               Strg_TO_Chars(Strg:= CONCAT_STRING(IN1 := #TMP_strTemp ,IN2 := DINT_TO_STRING(#IN_rgtStatusMarkers[#TMP_dMarkerIndex].dStatus)),
                         pChars:=#TMP_dIndex,
                         Cnt=>#TMP_uiNumChar,
                         Chars:=#AUX_rgcStatusTelegram);
               #TMP_dIndex+=#TMP_uiNumChar;

               #AUX_rgcStatusTelegram[#TMP_dIndex] := #STRSEPARATOR;
               #TMP_dIndex+=1;
           END_IF;

           IF (#IN_rgtStatusMarkers[#TMP_dMarkerIndex].dMarkerActualStatus <> #AUX_rgtStatusMarkers[#TMP_dMarkerIndex].dMarkerActualStatus) OR (#AUX_xResendAllStatus) THEN

               #AUX_rgtStatusMarkers[#TMP_dMarkerIndex].dMarkerActualStatus := #IN_rgtStatusMarkers[#TMP_dMarkerIndex].dMarkerActualStatus;        

               #TMP_strTemp := CONCAT_STRING(IN1 := #STRSTATUSMARKACTSTATUS ,IN2 := #TMP_strMarkerIndex);
               #TMP_strTemp := CONCAT_STRING(IN1 := #TMP_strTemp ,IN2 := '=');

               Strg_TO_Chars(Strg:= CONCAT_STRING(IN1 := #TMP_strTemp ,IN2 := DINT_TO_STRING(#IN_rgtStatusMarkers[#TMP_dMarkerIndex].dMarkerActualStatus)),
                         pChars:=#TMP_dIndex,
                         Cnt=>#TMP_uiNumChar,
                         Chars:=#AUX_rgcStatusTelegram);
               #TMP_dIndex+=#TMP_uiNumChar;

               #AUX_rgcStatusTelegram[#TMP_dIndex] := #STRSEPARATOR;
               #TMP_dIndex+=1;
           END_IF;*)


       END_FOR;

       END_REGION BPS_STATUS_TELEGRAM_MARKERS

       REGION BPS_STATUS_TELEGRAM_YCUTS

       FOR #TMP_dYCutIndex := 0 TO "DMAXYCUTBRIDGE_IND" DO

           #TMP_strYCutIndex := DINT_TO_STRING(#TMP_dYCutIndex + 1);   

           #TMP_strYCutIndex := DELETE(IN:=#TMP_strYCutIndex, L:=1, P:=1);

           //Prepare position information
           #TMP_strYCut := CONCAT_STRING(IN1 := #STRSTATUSYCUT ,IN2 := #TMP_strYCutIndex);

           IF (#IN_rgtStatusYCuts[#TMP_dYCutIndex].dBridgeStatus <> #AUX_rgtStatusYCuts[#TMP_dYCutIndex].dBridgeStatus) OR (#AUX_xResendAllStatus) THEN

               #AUX_rgtStatusYCuts[#TMP_dYCutIndex].dBridgeStatus := #IN_rgtStatusYCuts[#TMP_dYCutIndex].dBridgeStatus;        

               #TMP_strTemp := CONCAT_STRING(IN1 := #TMP_strYCut ,IN2 := #STRSTATUSYCUTSTATUS);

               Strg_TO_Chars(Strg:= CONCAT_STRING(IN1 := #TMP_strTemp ,IN2 := DINT_TO_STRING(#IN_rgtStatusYCuts[#TMP_dYCutIndex].dBridgeStatus)),
                         pChars:=#TMP_dIndex,
                         Cnt=>#TMP_uiNumChar,
                         Chars:=#AUX_rgcStatusTelegram);
               #TMP_dIndex+=#TMP_uiNumChar;

               #AUX_rgcStatusTelegram[#TMP_dIndex] := #STRSEPARATOR;
               #TMP_dIndex+=1;
           END_IF;

           IF (#IN_rgtStatusYCuts[#TMP_dYCutIndex].dDistanceSnapRoll_cmm <> #AUX_rgtStatusYCuts[#TMP_dYCutIndex].dDistanceSnapRoll_cmm) OR (#AUX_xResendAllStatus) THEN

               #AUX_rgtStatusYCuts[#TMP_dYCutIndex].dDistanceSnapRoll_cmm := #IN_rgtStatusYCuts[#TMP_dYCutIndex].dDistanceSnapRoll_cmm;        

               #TMP_strTemp := CONCAT_STRING(IN1 := #TMP_strYCut ,IN2 := #STRSTATUSYCUTSDISTSNAP);

               Strg_TO_Chars(Strg:= CONCAT_STRING(IN1 := #TMP_strTemp ,IN2 := DINT_TO_STRING(#IN_rgtStatusYCuts[#TMP_dYCutIndex].dDistanceSnapRoll_cmm)),
                         pChars:=#TMP_dIndex,
                         Cnt=>#TMP_uiNumChar,
                         Chars:=#AUX_rgcStatusTelegram);
               #TMP_dIndex+=#TMP_uiNumChar;

               #AUX_rgcStatusTelegram[#TMP_dIndex] := #STRSEPARATOR;
               #TMP_dIndex+=1;
           END_IF;


           FOR #TMP_dYCutHeadIndex := 0 TO "DMAXYHEADS_IND" DO

               #TMP_strHeadIndex := DINT_TO_STRING(#TMP_dYCutHeadIndex + 1);
               #TMP_strHeadIndex := DELETE(IN:=#TMP_strHeadIndex, L:= 1, P:=1);

               IF (#IN_rgtStatusYCuts[#TMP_dYCutIndex].rgdPosition_cmm[#TMP_dYCutHeadIndex] <> #AUX_rgtStatusYCuts[#TMP_dYCutIndex].rgdPosition_cmm[#TMP_dYCutHeadIndex]) OR (#AUX_xResendAllStatus) THEN

                   #AUX_rgtStatusYCuts[#TMP_dYCutIndex].rgdPosition_cmm[#TMP_dYCutHeadIndex] := #IN_rgtStatusYCuts[#TMP_dYCutIndex].rgdPosition_cmm[#TMP_dYCutHeadIndex];

                   #TMP_strTemp := CONCAT_STRING(IN1 := #TMP_strYCut ,IN2 := #STRSTATUSYCUTPOS);
                   #TMP_strTemp := CONCAT_STRING(IN1 := #TMP_strTemp, IN2 := #TMP_strHeadIndex);
                   #TMP_strTemp := CONCAT_STRING(IN1 := #TMP_strTemp,IN2 := '=');

                   Strg_TO_Chars(Strg:= CONCAT_STRING(IN1 := #TMP_strTemp ,IN2 := DINT_TO_STRING(#IN_rgtStatusYCuts[#TMP_dYCutIndex].rgdPosition_cmm[#TMP_dYCutHeadIndex])),
                         pChars:=#TMP_dIndex,
                         Cnt=>#TMP_uiNumChar,
                         Chars:=#AUX_rgcStatusTelegram);
                   #TMP_dIndex+=#TMP_uiNumChar;

                   #AUX_rgcStatusTelegram[#TMP_dIndex] := #STRSEPARATOR;
                   #TMP_dIndex+=1;
               END_IF;

               IF (#IN_rgtStatusYCuts[#TMP_dYCutIndex].rgxFireON[#TMP_dYCutHeadIndex] <> #AUX_rgtStatusYCuts[#TMP_dYCutIndex].rgxFireON[#TMP_dYCutHeadIndex]) OR (#AUX_xResendAllStatus) THEN

                   #AUX_rgtStatusYCuts[#TMP_dYCutIndex].rgxFireON[#TMP_dYCutHeadIndex] := #IN_rgtStatusYCuts[#TMP_dYCutIndex].rgxFireON[#TMP_dYCutHeadIndex];

                   #TMP_strTemp := CONCAT_STRING(IN1 := #TMP_strYCut ,IN2 := #STRSTATUSYCUTFIRE);
                   #TMP_strTemp := CONCAT_STRING(IN1 := #TMP_strTemp, IN2 := #TMP_strHeadIndex);
                   #TMP_strTemp := CONCAT_STRING(IN1 := #TMP_strTemp,IN2 := '=');

                   Strg_TO_Chars(Strg:= CONCAT_STRING(IN1 := #TMP_strTemp ,IN2 := DINT_TO_STRING(BOOL_TO_DINT(#IN_rgtStatusYCuts[#TMP_dYCutIndex].rgxFireON[#TMP_dYCutHeadIndex]))),
                         pChars:=#TMP_dIndex,
                         Cnt=>#TMP_uiNumChar,
                         Chars:=#AUX_rgcStatusTelegram);
                   #TMP_dIndex+=#TMP_uiNumChar;

                   #AUX_rgcStatusTelegram[#TMP_dIndex] := #STRSEPARATOR;
                   #TMP_dIndex+=1;
               END_IF;

               IF (#IN_rgtStatusYCuts[#TMP_dYCutIndex].rgxArmON[#TMP_dYCutHeadIndex] <> #AUX_rgtStatusYCuts[#TMP_dYCutIndex].rgxArmON[#TMP_dYCutHeadIndex]) OR (#AUX_xResendAllStatus) THEN

                   #AUX_rgtStatusYCuts[#TMP_dYCutIndex].rgxArmON[#TMP_dYCutHeadIndex] := #IN_rgtStatusYCuts[#TMP_dYCutIndex].rgxArmON[#TMP_dYCutHeadIndex];

                   #TMP_strTemp := CONCAT_STRING(IN1 := #TMP_strYCut ,IN2 := #STRSTATUSYCUTARM);
                   #TMP_strTemp := CONCAT_STRING(IN1 := #TMP_strTemp, IN2 := #TMP_strHeadIndex);
                   #TMP_strTemp := CONCAT_STRING(IN1 := #TMP_strTemp,IN2 := '=');

                   Strg_TO_Chars(Strg:= CONCAT_STRING(IN1 := #TMP_strTemp ,IN2 := DINT_TO_STRING(BOOL_TO_DINT(#IN_rgtStatusYCuts[#TMP_dYCutIndex].rgxArmON[#TMP_dYCutHeadIndex]))),
                         pChars:=#TMP_dIndex,
                         Cnt=>#TMP_uiNumChar,
                         Chars:=#AUX_rgcStatusTelegram);
                   #TMP_dIndex+=#TMP_uiNumChar;

                   #AUX_rgcStatusTelegram[#TMP_dIndex] := #STRSEPARATOR;
                   #TMP_dIndex+=1;
               END_IF;

               IF (#IN_rgtStatusYCuts[#TMP_dYCutIndex].rgxHeadProdOn[#TMP_dYCutHeadIndex] <> #AUX_rgtStatusYCuts[#TMP_dYCutIndex].rgxHeadProdOn[#TMP_dYCutHeadIndex]) OR (#AUX_xResendAllStatus) THEN

                   #AUX_rgtStatusYCuts[#TMP_dYCutIndex].rgxHeadProdOn[#TMP_dYCutHeadIndex] := #IN_rgtStatusYCuts[#TMP_dYCutIndex].rgxHeadProdOn[#TMP_dYCutHeadIndex];

                   #TMP_strTemp := CONCAT_STRING(IN1 := #TMP_strYCut ,IN2 := #STRSTATUSYCUTPROD);
                   #TMP_strTemp := CONCAT_STRING(IN1 := #TMP_strTemp, IN2 := #TMP_strHeadIndex);
                   #TMP_strTemp := CONCAT_STRING(IN1 := #TMP_strTemp,IN2 := '=');

                   Strg_TO_Chars(Strg:= CONCAT_STRING(IN1 := #TMP_strTemp ,IN2 := DINT_TO_STRING(BOOL_TO_DINT(#IN_rgtStatusYCuts[#TMP_dYCutIndex].rgxHeadProdOn[#TMP_dYCutHeadIndex]))),
                         pChars:=#TMP_dIndex,
                         Cnt=>#TMP_uiNumChar,
                         Chars:=#AUX_rgcStatusTelegram);
                   #TMP_dIndex+=#TMP_uiNumChar;

                   #AUX_rgcStatusTelegram[#TMP_dIndex] := #STRSEPARATOR;
                   #TMP_dIndex+=1;
               END_IF;

           END_FOR;


       END_FOR;

      // #AUX_xResendAllStatus := FALSE;


       END_REGION BPS_STATUS_TELEGRAM_YCUTS


       #AUX_rgcStatusTelegram[#TMP_dIndex] := #STR_CR;
       #TMP_dIndex+=1;

       #AUX_rgcStatusTelegram[#TMP_dIndex] := #STR_LF;

       #AUX_dStatusTelegramNumByte := #TMP_dIndex + 1;

       IF #AUX_dStatusTelegramCounter >= #DMAXTELEGRAMCOUNTER THEN
           #AUX_dStatusTelegramCounter := 1;
       ELSE
           #AUX_dStatusTelegramCounter += 1;
       END_IF;

       IF (((#IN_xBPSServerA) AND (#IN_tStatusGeneral.dExtOptSelected = 1)) OR
           ((NOT #IN_xBPSServerA) AND (#IN_tStatusGeneral.dExtOptSelected = 2))) THEN

           IF #AUX_dStatusServerCounter >= #DMAXTELEGRAMCOUNTER THEN
               #AUX_dStatusServerCounter := 1;
           ELSE
               #AUX_dStatusServerCounter += 1;
           END_IF;

       END_IF;    
       #ST_xStatusTelegramAvail := TRUE;

   END_IF;





   END_REGION BPS_STATUS_TELEGRAM

   REGION BPS_SEND_INFORMATION

   //Initialize connection data in case of reset
   IF #IN_xGeneralReset THEN

       #AUX_tConnData.InterfaceId := #IN_tInterfaceID;
       #AUX_tConnData.ID := #IN_tID;
       #AUX_tConnData.ConnectionType := #BCONNTYPE;
       #AUX_tConnData.ActiveEstablished := TRUE;
       #AUX_tConnData.RemoteAddress := #IN_tRemoteAddress;
       #AUX_tConnData.RemotePort := #IN_uiRemotePort;
       #AUX_tConnData.LocalPort := 0;

       //Reset della fasi
       #TMP_dwValue := 0;
       SCATTER(IN:=#TMP_dwValue,
               OUT=>#tPhasesNetwork);

       //Reset others data
       #ST_xRetrySendTelegram := FALSE;
       #AUX_dSendTelegramNumByte := 0;
       #TMP_cValue := ' ';

       FILL_BLK(IN:=#TMP_cValue,
                COUNT:=DINT_TO_ULINT(#DSENDTELEGRAMSIZE),
                OUT=>#AUX_rgcSendTelegram[0]);


   END_IF;

   #AUX_xResetSendConnection := #IN_xGeneralReset OR (#FB_TSend.s_TDIAG_Status.State <> b#16#04 AND #IN_xResetAlarms);


   IF NOT #ST_xPhasesInProgress AND #IN_xThisPLCActive AND
           (#ST_xPlateTelegramAvail OR 
           #ST_xStatusTelegramAvail OR 
           #ST_xDefectTelegramAvail OR 
           #ST_xRibbonTelegramAvail OR 
           #ST_xEventsTelegramAvail OR
           #ST_xRibbonTelegramAvail OR 
           #ST_xRetrySendTelegram) THEN

       IF NOT #ST_xRetrySendTelegram THEN

           //Fill the send buffer with the status telegram and plate
           #AUX_dSendTelegramNumByte := 0;

           IF #ST_xPlateTelegramAvail THEN

               MOVE_BLK(IN:=#AUX_rgcPlateTelegram[0],
                        COUNT:=DINT_TO_ULINT(#AUX_dPlateTelegramNumByte),
                        OUT=>#AUX_rgcSendTelegram[0]);

               #AUX_dSendTelegramNumByte:= #AUX_dPlateTelegramNumByte;

               #ST_xPlateTelegramAvail := FALSE;
               #AUX_xResendAllPlate := FALSE;
           ELSIF #ST_xStatusTelegramAvail THEN

               MOVE_BLK(IN := #AUX_rgcStatusTelegram[0],
                        COUNT := DINT_TO_ULINT(#AUX_dStatusTelegramNumByte),
                        OUT => #AUX_rgcSendTelegram[0]);

               #AUX_dSendTelegramNumByte := #AUX_dStatusTelegramNumByte;

               #ST_xStatusTelegramAvail := FALSE;
               #AUX_xResendAllStatus := FALSE;


           ELSIF #ST_xDefectTelegramAvail THEN

               MOVE_BLK(IN:=#AUX_rgcDefectTelegram[0],
                        COUNT:=DINT_TO_ULINT(#AUX_dDefectTelegramNumByte),
                        OUT=>#AUX_rgcSendTelegram[0]);

               #AUX_dSendTelegramNumByte:= #AUX_dDefectTelegramNumByte;

               #ST_xDefectTelegramAvail := FALSE;

           ELSIF #ST_xEventsTelegramAvail THEN

               MOVE_BLK(IN:=#AUX_rgcEventsTelegram[0],
                        COUNT:=DINT_TO_ULINT(#AUX_dEventsTelegramNumByte),
                        OUT=>#AUX_rgcSendTelegram[0]);

               #AUX_dSendTelegramNumByte:= #AUX_dEventsTelegramNumByte;

               #ST_xEventsTelegramAvail := FALSE;

           ELSIF #ST_xRibbonTelegramAvail THEN

               MOVE_BLK(IN:=#AUX_rgcRibbonTelegram[0],
                        COUNT:=DINT_TO_ULINT(#AUX_dRibbonTelegramNumByte),
                        OUT=>#AUX_rgcSendTelegram[0]);

               #AUX_dSendTelegramNumByte:= #AUX_dRibbonTelegramNumByte;

               #ST_xRibbonTelegramAvail := FALSE;

          ELSIF #ST_xStatusTelegramAvail THEN

               MOVE_BLK(IN:=#AUX_rgcStatusTelegram[0],
                        COUNT:=DINT_TO_ULINT(#AUX_dStatusTelegramNumByte),
                        OUT=>#AUX_rgcSendTelegram[0]);

               #AUX_dSendTelegramNumByte:= #AUX_dStatusTelegramNumByte;

               #ST_xStatusTelegramAvail := FALSE;
               #AUX_xResendAllStatus := FALSE;
           END_IF;

       END_IF;


       #tPhasesNetwork.xSendBufferInProgress := TRUE; 

   END_IF;


   #FB_TSend(REQ:=#tPhasesNetwork.xSendBufferInProgress,
             CONT:=#IN_xThisPLCActive,
             LEN:=DINT_TO_UDINT(#AUX_dSendTelegramNumByte),
             CONNECT:=#AUX_tConnData,
             DATA:=#AUX_rgcSendTelegram,
             COM_RST:=#AUX_xResetSendConnection);


   //Manage send feedback
   IF #tPhasesNetwork.xSendBufferInProgress AND 
                                           (#FB_TSend.DONE OR
                                           #FB_TSend.ERROR OR 
                                           NOT #FB_TSend.BUSY) THEN

       #tPhasesNetwork.xSendBufferInProgress := FALSE;
       #tPhasesNetwork.xEndSendBufferInProgress := TRUE;
       #ST_xRetrySendTelegram := FALSE;
       IF NOT #FB_TSend.DONE THEN

           #ST_xRetrySendTelegram := TRUE;

       END_IF;

   ELSE

       #tPhasesNetwork.xEndSendBufferInProgress := FALSE;
   END_IF;

   //Calculate phase in progress
   GATHER(IN:=#tPhasesNetwork,
          OUT=>#TMP_dwValue);

   IF #TMP_dwValue <> 0 THEN
       #ST_xPhasesInProgress := TRUE;
   ELSE
       #ST_xPhasesInProgress := FALSE;
   END_IF;




   END_REGION BPS_SEND_INFORMATION

   REGION BPS_RECEIVE_INFORMATION

   #FB_TRecv(EN_R:=#IN_xThisPLCActive,
             CONT:=#IN_xThisPLCActive,
             LEN:=0,
             ADHOC:=TRUE,
             CONNECT:=#AUX_tConnData,
             DATA:=#AUX_rgcRecvTelegram,
             COM_RST:=#AUX_xResetSendConnection);

   IF #FB_TRecv.DONE THEN

       IF (#FB_TRecv.RCVD_LEN > 0) AND (UDINT_TO_DINT(#FB_TRecv.RCVD_LEN) + #AUX_dNumByteRecvBuffer < #DRECVBUFFERSIZE) THEN

           //Copy the received data
           #TMP_iRetVal := MOVE_BLK_VARIANT(SRC:=#AUX_rgcRecvTelegram, COUNT:=#FB_TRecv.RCVD_LEN, SRC_INDEX:=0, DEST_INDEX:=#AUX_dNumByteRecvBuffer, DEST=>#AUX_rgcRecvBuffer);
           #AUX_dNumByteRecvBuffer += UDINT_TO_DINT(#FB_TRecv.RCVD_LEN);

       END_IF;

   END_IF;

   //Analyze telegrams 
   FOR #TMP_dIndex := 0 TO #AUX_dNumByteRecvBuffer - 2 DO

       IF (#AUX_rgcRecvBuffer[#TMP_dIndex] = #STR_CR) AND (#AUX_rgcRecvBuffer[#TMP_dIndex + 1] = #STR_LF) THEN

           //End of packet found. Move the data to a string
           #TMP_iRetVal := MOVE_BLK_VARIANT(SRC:=#AUX_rgcRecvBuffer, COUNT:= DINT_TO_UDINT(#TMP_dIndex) + 2 , SRC_INDEX:= 0, DEST_INDEX:= 0, DEST=>#AUX_rgcAnalyzedTelegram);

           IF (#TMP_dIndex + 2) < #AUX_dNumByteRecvBuffer THEN
               #TMP_iRetVal := MOVE_BLK_VARIANT(SRC:=#AUX_rgcRecvBuffer, COUNT:=DINT_TO_UDINT(#AUX_dNumByteRecvBuffer - (#TMP_dIndex + 2))   , SRC_INDEX:= #TMP_dIndex + 2 , DEST_INDEX:= 0, DEST=>#AUX_rgcRecvBuffer);
           ELSE
               #AUX_dNumByteRecvBuffer := 0;
           END_IF;
           #TMP_udCountString := 0;
           #TMP_udPosition := 0;
           #TMP_cSeparator := #STRSEPARATOR;

           #TMP_cEndSeparator := #STR_LF;
           //Split the telegram and manage it
           #TMP_iRetVal := SPLIT(Mode:=0, RecSeparator:=#TMP_cSeparator, EndSeparator:=#TMP_cEndSeparator, SrcArray:=#AUX_rgcAnalyzedTelegram, Count=>#TMP_udCountString, DstStruct:=#AUX_rgstrMessageString, Position:=#TMP_udPosition);

   REGION BPS_RECEIVE_EVENT 
           //Check the received message 'D'
           IF (#AUX_rgstrMessageString[0] = CHAR_TO_STRING(#STREVENTSTELEGRAMID)) AND (#TMP_udCountString = 16) THEN

               //Event code
               #TMP_cSeparator := '=';
               #TMP_uiCount := 0;


               Strg_TO_Chars(Strg:=#AUX_rgstrMessageString[2],
                             pChars:=0,
                             Cnt=>#TMP_uiCount,
                             Chars:=#AUX_rgcMetaData);
               #AUX_rgcMetaData[#TMP_uiCount] := #STR_LF;
               #TMP_udPosition := 0;
               #TMP_iRetVal := SPLIT(  Mode:=0, 
                                       RecSeparator:=#TMP_cSeparator, 
                                       EndSeparator:=#TMP_cEndSeparator, 
                                       SrcArray:=#AUX_rgcMetaData, 
                                       Count=>#TMP_udCountString, 
                                       DstStruct:=#AUX_rgstrSingleMexString, 
                                       Position:=#TMP_udPosition);
               IF ( #TMP_udCountString = 2) AND #AUX_rgstrSingleMexString[0] = 'Cd' THEN
                   #AUX_tRecvMessage.dCodeEvent := STRING_TO_DINT(#AUX_rgstrSingleMexString[1]);
               ELSE 
                   #AUX_tRecvMessage.dCodeEvent := 0;
               END_IF;

               //Ident
               #TMP_cSeparator := '=';
               #TMP_uiCount := 0;
               Strg_TO_Chars(Strg:=#AUX_rgstrMessageString[4],
                             pChars:=0,
                             Cnt=>#TMP_uiCount,
                             Chars:=#AUX_rgcMetaData);
               #AUX_rgcMetaData[#TMP_uiCount] := #STR_LF;
               #TMP_udPosition := 0;
               #TMP_iRetVal := SPLIT(  Mode:=0, 
                                       RecSeparator:=#TMP_cSeparator, 
                                       EndSeparator:=#TMP_cEndSeparator, 
                                       SrcArray:=#AUX_rgcMetaData, 
                                       Count=>#TMP_udCountString, 
                                       DstStruct:=#AUX_rgstrSingleMexString, 
                                       Position:=#TMP_udPosition);
               IF ( #TMP_udCountString = 2) AND #AUX_rgstrSingleMexString[0] = 'Id' THEN
                   #AUX_tRecvMessage.strIdent := #AUX_rgstrSingleMexString[1];
               ELSE 
                   #AUX_tRecvMessage.strIdent := '';
               END_IF;

               //Data 1
               #TMP_cSeparator := '=';
               #TMP_uiCount := 0;
               Strg_TO_Chars(Strg:=#AUX_rgstrMessageString[5],
                             pChars:=0,
                             Cnt=>#TMP_uiCount,
                             Chars:=#AUX_rgcMetaData);
               #AUX_rgcMetaData[#TMP_uiCount] := #STR_LF;
               #TMP_udPosition := 0;
               #TMP_iRetVal := SPLIT(  Mode:=0, 
                                       RecSeparator:=#TMP_cSeparator, 
                                       EndSeparator:=#TMP_cEndSeparator, 
                                       SrcArray:=#AUX_rgcMetaData, 
                                       Count=>#TMP_udCountString, 
                                       DstStruct:=#AUX_rgstrSingleMexString, 
                                       Position:=#TMP_udPosition);
               IF ( #TMP_udCountString = 2) AND #AUX_rgstrSingleMexString[0] = 'D1' THEN
                   #AUX_tRecvMessage.dEvent1 := STRING_TO_DINT(#AUX_rgstrSingleMexString[1]);
               ELSE 
                   #AUX_tRecvMessage.dEvent1 := 0;
               END_IF;

               //Data 2
               #TMP_cSeparator := '=';
               #TMP_uiCount := 0;
               Strg_TO_Chars(Strg:=#AUX_rgstrMessageString[6],
                             pChars:=0,
                             Cnt=>#TMP_uiCount,
                             Chars:=#AUX_rgcMetaData);
               #AUX_rgcMetaData[#TMP_uiCount] := #STR_LF;
               #TMP_udPosition := 0;
               #TMP_iRetVal := SPLIT(  Mode:=0, 
                                       RecSeparator:=#TMP_cSeparator, 
                                       EndSeparator:=#TMP_cEndSeparator, 
                                       SrcArray:=#AUX_rgcMetaData, 
                                       Count=>#TMP_udCountString, 
                                       DstStruct:=#AUX_rgstrSingleMexString, 
                                       Position:=#TMP_udPosition);
               IF ( #TMP_udCountString = 2) AND #AUX_rgstrSingleMexString[0] = 'D2' THEN
                   #AUX_tRecvMessage.dEvent2 := STRING_TO_DINT(#AUX_rgstrSingleMexString[1]);
               ELSE 
                   #AUX_tRecvMessage.dEvent2 := 0;
               END_IF;

               //Data 3
               #TMP_cSeparator := '=';
               #TMP_uiCount := 0;
               Strg_TO_Chars(Strg:=#AUX_rgstrMessageString[7],
                             pChars:=0,
                             Cnt=>#TMP_uiCount,
                             Chars:=#AUX_rgcMetaData);
               #AUX_rgcMetaData[#TMP_uiCount] := #STR_LF;
               #TMP_udPosition := 0;
               #TMP_iRetVal := SPLIT(  Mode:=0, 
                                       RecSeparator:=#TMP_cSeparator, 
                                       EndSeparator:=#TMP_cEndSeparator, 
                                       SrcArray:=#AUX_rgcMetaData, 
                                       Count=>#TMP_udCountString, 
                                       DstStruct:=#AUX_rgstrSingleMexString, 
                                       Position:=#TMP_udPosition);
               IF ( #TMP_udCountString = 2) AND #AUX_rgstrSingleMexString[0] = 'D3' THEN
                   #AUX_tRecvMessage.dEvent3 := STRING_TO_DINT(#AUX_rgstrSingleMexString[1]);
               ELSE 
                   #AUX_tRecvMessage.dEvent3 := 0;
               END_IF;

               //Data 4
               #TMP_cSeparator := '=';
               #TMP_uiCount := 0;
               Strg_TO_Chars(Strg:=#AUX_rgstrMessageString[8],
                             pChars:=0,
                             Cnt=>#TMP_uiCount,
                             Chars:=#AUX_rgcMetaData);
               #AUX_rgcMetaData[#TMP_uiCount] := #STR_LF;
               #TMP_udPosition := 0;
               #TMP_iRetVal := SPLIT(  Mode:=0, 
                                       RecSeparator:=#TMP_cSeparator, 
                                       EndSeparator:=#TMP_cEndSeparator, 
                                       SrcArray:=#AUX_rgcMetaData, 
                                       Count=>#TMP_udCountString, 
                                       DstStruct:=#AUX_rgstrSingleMexString, 
                                       Position:=#TMP_udPosition);
               IF ( #TMP_udCountString = 2) AND #AUX_rgstrSingleMexString[0] = 'D4' THEN
                   #AUX_tRecvMessage.dEvent4 := STRING_TO_DINT(#AUX_rgstrSingleMexString[1]);
               ELSE 
                   #AUX_tRecvMessage.dEvent4 := 0;
               END_IF;

               //Data 5
               #TMP_cSeparator := '=';
               #TMP_uiCount := 0;
               Strg_TO_Chars(Strg:=#AUX_rgstrMessageString[9],
                             pChars:=0,
                             Cnt=>#TMP_uiCount,
                             Chars:=#AUX_rgcMetaData);
               #AUX_rgcMetaData[#TMP_uiCount] := #STR_LF;
               #TMP_udPosition := 0;
               #TMP_iRetVal := SPLIT(  Mode:=0, 
                                       RecSeparator:=#TMP_cSeparator, 
                                       EndSeparator:=#TMP_cEndSeparator, 
                                       SrcArray:=#AUX_rgcMetaData, 
                                       Count=>#TMP_udCountString, 
                                       DstStruct:=#AUX_rgstrSingleMexString, 
                                       Position:=#TMP_udPosition);
               IF ( #TMP_udCountString = 2) AND #AUX_rgstrSingleMexString[0] = 'D5' THEN
                   #AUX_tRecvMessage.dEvent5 := STRING_TO_DINT(#AUX_rgstrSingleMexString[1]);
               ELSE 
                   #AUX_tRecvMessage.dEvent5 := 0;
               END_IF;

               //Data 6
               #TMP_cSeparator := '=';
               #TMP_uiCount := 0;
               Strg_TO_Chars(Strg:=#AUX_rgstrMessageString[10],
                             pChars:=0,
                             Cnt=>#TMP_uiCount,
                             Chars:=#AUX_rgcMetaData);
               #AUX_rgcMetaData[#TMP_uiCount] := #STR_LF;
               #TMP_udPosition := 0;
               #TMP_iRetVal := SPLIT(  Mode:=0, 
                                       RecSeparator:=#TMP_cSeparator, 
                                       EndSeparator:=#TMP_cEndSeparator, 
                                       SrcArray:=#AUX_rgcMetaData, 
                                       Count=>#TMP_udCountString, 
                                       DstStruct:=#AUX_rgstrSingleMexString, 
                                       Position:=#TMP_udPosition);
               IF ( #TMP_udCountString = 2) AND #AUX_rgstrSingleMexString[0] = 'D6' THEN
                   #AUX_tRecvMessage.dEvent6 := STRING_TO_DINT(#AUX_rgstrSingleMexString[1]);
               ELSE 
                   #AUX_tRecvMessage.dEvent6 := 0;
               END_IF;

               //Data 7
               #TMP_cSeparator := '=';
               #TMP_uiCount := 0;
               Strg_TO_Chars(Strg:=#AUX_rgstrMessageString[11],
                             pChars:=0,
                             Cnt=>#TMP_uiCount,
                             Chars:=#AUX_rgcMetaData);
               #AUX_rgcMetaData[#TMP_uiCount] := #STR_LF;
               #TMP_udPosition := 0;
               #TMP_iRetVal := SPLIT(  Mode:=0, 
                                       RecSeparator:=#TMP_cSeparator, 
                                       EndSeparator:=#TMP_cEndSeparator, 
                                       SrcArray:=#AUX_rgcMetaData, 
                                       Count=>#TMP_udCountString, 
                                       DstStruct:=#AUX_rgstrSingleMexString, 
                                       Position:=#TMP_udPosition);
               IF ( #TMP_udCountString = 2) AND #AUX_rgstrSingleMexString[0] = 'D7' THEN
                   #AUX_tRecvMessage.dEvent7 := STRING_TO_DINT(#AUX_rgstrSingleMexString[1]);
               ELSE 
                   #AUX_tRecvMessage.dEvent7 := 0;
               END_IF;

               //Data 8
               #TMP_cSeparator := '=';
               #TMP_uiCount := 0;
               Strg_TO_Chars(Strg:=#AUX_rgstrMessageString[12],
                             pChars:=0,
                             Cnt=>#TMP_uiCount,
                             Chars:=#AUX_rgcMetaData);
               #AUX_rgcMetaData[#TMP_uiCount] := #STR_LF;
               #TMP_udPosition := 0;
               #TMP_iRetVal := SPLIT(  Mode:=0, 
                                       RecSeparator:=#TMP_cSeparator, 
                                       EndSeparator:=#TMP_cEndSeparator, 
                                       SrcArray:=#AUX_rgcMetaData, 
                                       Count=>#TMP_udCountString, 
                                       DstStruct:=#AUX_rgstrSingleMexString, 
                                       Position:=#TMP_udPosition);
               IF ( #TMP_udCountString = 2) AND #AUX_rgstrSingleMexString[0] = 'D8' THEN
                   #AUX_tRecvMessage.dEvent8 := STRING_TO_DINT(#AUX_rgstrSingleMexString[1]);
               ELSE 
                   #AUX_tRecvMessage.dEvent8 := 0;
               END_IF;

               //Data 9
               #TMP_cSeparator := '=';
               #TMP_uiCount := 0;
               Strg_TO_Chars(Strg:=#AUX_rgstrMessageString[13],
                             pChars:=0,
                             Cnt=>#TMP_uiCount,
                             Chars:=#AUX_rgcMetaData);
               #AUX_rgcMetaData[#TMP_uiCount] := #STR_LF;
               #TMP_udPosition := 0;
               #TMP_iRetVal := SPLIT(  Mode:=0, 
                                       RecSeparator:=#TMP_cSeparator, 
                                       EndSeparator:=#TMP_cEndSeparator, 
                                       SrcArray:=#AUX_rgcMetaData, 
                                       Count=>#TMP_udCountString, 
                                       DstStruct:=#AUX_rgstrSingleMexString, 
                                       Position:=#TMP_udPosition);
               IF ( #TMP_udCountString = 2) AND #AUX_rgstrSingleMexString[0] = 'D9' THEN
                   #AUX_tRecvMessage.dEvent9 := STRING_TO_DINT(#AUX_rgstrSingleMexString[1]);
               ELSE 
                   #AUX_tRecvMessage.dEvent9 := 0;
               END_IF;

               //Data 10
               #TMP_cSeparator := '=';
               #TMP_uiCount := 0;
               Strg_TO_Chars(Strg:=#AUX_rgstrMessageString[14],
                             pChars:=0,
                             Cnt=>#TMP_uiCount,
                             Chars:=#AUX_rgcMetaData);
               #AUX_rgcMetaData[#TMP_uiCount] := #STR_LF;
               #TMP_udPosition := 0;
               #TMP_iRetVal := SPLIT(  Mode:=0, 
                                       RecSeparator:=#TMP_cSeparator, 
                                       EndSeparator:=#TMP_cEndSeparator, 
                                       SrcArray:=#AUX_rgcMetaData, 
                                       Count=>#TMP_udCountString, 
                                       DstStruct:=#AUX_rgstrSingleMexString, 
                                       Position:=#TMP_udPosition);
               IF ( #TMP_udCountString = 2) AND #AUX_rgstrSingleMexString[0] = 'D10' THEN
                   #AUX_tRecvMessage.dEvent10 := STRING_TO_DINT(#AUX_rgstrSingleMexString[1]);
               ELSE 
                   #AUX_tRecvMessage.dEvent10 := 0;
               END_IF;

               "RP_AddMessageV2"(IN_xInit:=FALSE,
                                 IN_dCodeEvent:=#AUX_tRecvMessage.dCodeEvent,
                                 IN_strIndet_Max4Chars:=#AUX_tRecvMessage.strIdent,
                                 IN_dValue1:=#AUX_tRecvMessage.dEvent1,
                                 IN_dValue2:=#AUX_tRecvMessage.dEvent2,
                                 IN_dValue3:=#AUX_tRecvMessage.dEvent3,
                                 IN_dValue4:=#AUX_tRecvMessage.dEvent4,
                                 IN_dValue5:=#AUX_tRecvMessage.dEvent5,
                                 IN_dValue6:=#AUX_tRecvMessage.dEvent6,
                                 IN_dValue7:=#AUX_tRecvMessage.dEvent7,
                                 IN_dValue8:=#AUX_tRecvMessage.dEvent8,
                                 IN_dValue9:=#AUX_tRecvMessage.dEvent9,
                                 IN_dValue10:=#AUX_tRecvMessage.dEvent10,
                                 INO_tBuffer:=#INO_tAddMessageFromOpt,
                                 INO_xError:=#INO_xMessageAnomaly);

           END_IF;
   END_REGION BPS_RECEIVE_EVENT 

       END_IF;

   END_FOR;  





   END_REGION BPS_RECEIVE_INFORMATION
END_FUNCTION_BLOCK

// folder: 03_Programs_Logics/MCC1200/15_ColdBackup

FUNCTION_BLOCK "FB_ColdBackupManager_V1.00"   // FB14, LAD
{ S7_Optimized_Access := 'TRUE' }
VERSION : 0.1
   VAR_INPUT
      IN_xGeneralReset : Bool;   // General reset
      IN_xResetAlarms : Bool;   // Reset alarms
      IN_tHWInterface : Hw_Interface;   // HW interface id
      IN_tConfDataMaster : Struct   // Configuration data master CPU
         Header : IF_CONF_Header;
         IPData : IF_CONF_v4;
         NoS : IF_CONF_NOS;
         NTP : IF_CONF_NTP;
         IP_V6 : IF_CONF_v6;
         MAC : IF_CONF_MAC;
         DNS : IF_CONF_DNS;
      END_STRUCT;
      IN_tConfDataBackup : Struct   // Configuration data backup CPU
         Header : IF_CONF_Header;
         IPData : IF_CONF_v4;
         NoS : IF_CONF_NOS;
         NTP : IF_CONF_NTP;
         IP_V6 : IF_CONF_v6;
         MAC : IF_CONF_MAC;
         DNS : IF_CONF_DNS;
      END_STRUCT;
      IN_xThisPLCActive : Bool;   // This PLC Active
   END_VAR
   VAR RETAIN
      tHMR : Struct
         dSpare : DInt;
      END_STRUCT;
      tHMW : Struct
         dSpare : DInt;
      END_STRUCT;
   END_VAR
   VAR
      tALM : Struct   // HMI Alarms
         tS : Struct   // Stopping faults
            xSpare_0 : Bool;
            xSpare_1 : Bool;
            xSpare_2 : Bool;
            xSpare_3 : Bool;
            xSpare_4 : Bool;
            xSpare_5 : Bool;
            xSpare_6 : Bool;
            xSpare_7 : Bool;
            xSpare_8 : Bool;
            xSpare_9 : Bool;
            xSpare_10 : Bool;
            xSpare_11 : Bool;
            xSpare_12 : Bool;
            xSpare_13 : Bool;
            xSpare_14 : Bool;
            xSpare_15 : Bool;
            xSpare_16 : Bool;
            xSpare_17 : Bool;
            xSpare_18 : Bool;
            xSpare_19 : Bool;
            xSpare_20 : Bool;
            xSpare_21 : Bool;
            xSpare_22 : Bool;
            xSpare_23 : Bool;
            xSpare_24 : Bool;
            xSpare_25 : Bool;
            xSpare_26 : Bool;
            xSpare_27 : Bool;
            xSpare_28 : Bool;
            xSpare_29 : Bool;
            xSpare_30 : Bool;
            xSpare_31 : Bool;
         END_STRUCT;
         tF : Struct   // Faults
            xSpare_0 : Bool;
            xSpare_1 : Bool;
            xSpare_2 : Bool;
            xSpare_3 : Bool;
            xSpare_4 : Bool;
            xSpare_5 : Bool;
            xSpare_6 : Bool;
            xSpare_7 : Bool;
            xSpare_8 : Bool;
            xSpare_9 : Bool;
            xSpare_10 : Bool;
            xSpare_11 : Bool;
            xSpare_12 : Bool;
            xSpare_13 : Bool;
            xSpare_14 : Bool;
            xSpare_15 : Bool;
            xSpare_16 : Bool;
            xSpare_17 : Bool;
            xSpare_18 : Bool;
            xSpare_19 : Bool;
            xSpare_20 : Bool;
            xSpare_21 : Bool;
            xSpare_22 : Bool;
            xSpare_23 : Bool;
            xSpare_24 : Bool;
            xSpare_25 : Bool;
            xSpare_26 : Bool;
            xSpare_27 : Bool;
            xSpare_28 : Bool;
            xSpare_29 : Bool;
            xSpare_30 : Bool;
            xSpare_31 : Bool;
         END_STRUCT;
         tW : Struct   // Warnings
            xSpare_0 : Bool;
            xSpare_1 : Bool;
            xSpare_2 : Bool;
            xSpare_3 : Bool;
            xSpare_4 : Bool;
            xSpare_5 : Bool;
            xSpare_6 : Bool;
            xSpare_7 : Bool;
            xSpare_8 : Bool;
            xSpare_9 : Bool;
            xSpare_10 : Bool;
            xSpare_11 : Bool;
            xSpare_12 : Bool;
            xSpare_13 : Bool;
            xSpare_14 : Bool;
            xSpare_15 : Bool;
            xSpare_16 : Bool;
            xSpare_17 : Bool;
            xSpare_18 : Bool;
            xSpare_19 : Bool;
            xSpare_20 : Bool;
            xSpare_21 : Bool;
            xSpare_22 : Bool;
            xSpare_23 : Bool;
            xSpare_24 : Bool;
            xSpare_25 : Bool;
            xSpare_26 : Bool;
            xSpare_27 : Bool;
            xSpare_28 : Bool;
            xSpare_29 : Bool;
            xSpare_30 : Bool;
            xSpare_31 : Bool;
         END_STRUCT;
      END_STRUCT;
      STC_OSR_xThisPLCBackup : Bool;   // OSR This PLC backup
      STC_OSR_xThisPLCActive : Bool;   // OSR This PLC active
      STC_ST_xRequestIpConfig : Bool;   // IP configuration request
      FB_T_Config : T_CONFIG;   // FB T config istance
      STC_tConfData : Struct
         Header : IF_CONF_Header;
         IPData : IF_CONF_v4;
         NoS : IF_CONF_NOS;
         NTP : IF_CONF_NTP;
         IP_V6 : IF_CONF_v6;
         MAC : IF_CONF_MAC;
         DNS : IF_CONF_DNS;
      END_STRUCT;
   END_VAR
   VAR_TEMP   // added for the SCL form of the ladder/FBD networks
      _w1 : Bool;
      _w2 : Bool;
   END_VAR
BEGIN

REGION Network 1: ####_COSTANTS_####
END_REGION

REGION Network 2: ####_MATCH_####
END_REGION

REGION Network 3: ####_ALARMS_####
END_REGION

REGION Network 4: ####_HMI_LOGICS_####
END_REGION

REGION Network 5: ####_STATUSES_####
END_REGION

REGION Network 6: ####_PHASES_&_LOGICS_####
END_REGION

REGION Network 7: IP configuration request
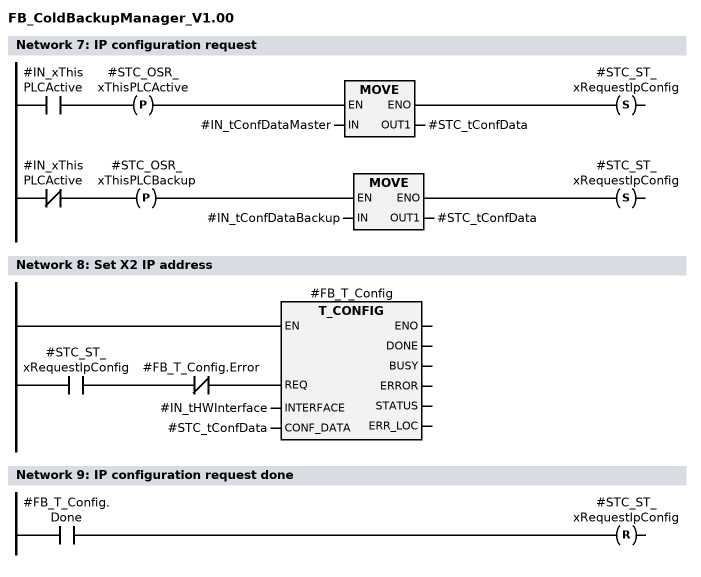
   RUNG wire#powerrail
      Contact( #IN_xThisPLCActive )
      P_Trig( #STC_OSR_xThisPLCActive )
      Move(in := #IN_tConfDataMaster, out1 => #STC_tConfData)
      S_Coil( #STC_ST_xRequestIpConfig )
   END_RUNG
   RUNG wire#powerrail
      I_Contact( #IN_xThisPLCActive )
      P_Trig( #STC_OSR_xThisPLCBackup )
      Move(in := #IN_tConfDataBackup, out1 => #STC_tConfData)
      S_Coil( #STC_ST_xRequestIpConfig )
   END_RUNG
   // the same network as SCL:
   #_w1 := #IN_xThisPLCActive AND NOT #STC_OSR_xThisPLCActive;   // rising edge
   #STC_OSR_xThisPLCActive := #IN_xThisPLCActive;
   IF #_w1 THEN
       #STC_tConfData := #IN_tConfDataMaster;
       #STC_ST_xRequestIpConfig := TRUE;
   END_IF;
   #_w2 := NOT #IN_xThisPLCActive AND NOT #STC_OSR_xThisPLCBackup;   // rising edge
   #STC_OSR_xThisPLCBackup := NOT #IN_xThisPLCActive;
   IF #_w2 THEN
       #STC_tConfData := #IN_tConfDataBackup;
       #STC_ST_xRequestIpConfig := TRUE;
   END_IF;
END_REGION

REGION Network 8: Set X2 IP address
   #FB_T_Config(Req := #STC_ST_xRequestIpConfig AND NOT #FB_T_Config.Error,   // T_CONFIG
                Interface := #IN_tHWInterface,
                Conf_Data := #STC_tConfData);
END_REGION

REGION Network 9: IP configuration request done
   RUNG wire#powerrail
      Contact( #FB_T_Config.Done )
      R_Coil( #STC_ST_xRequestIpConfig )
   END_RUNG
   // the same network as SCL:
   IF #FB_T_Config.Done THEN #STC_ST_xRequestIpConfig := FALSE; END_IF;
END_REGION

REGION Network 10 (SCL): ####_HMI_STATUSES_####
END_REGION

REGION Network 11: ####_OUTPUTS_####
END_REGION
END_FUNCTION_BLOCK

FUNCTION_BLOCK "FB_SwhitcTxRxColdBack_V1.00"   // FB27, LAD
{ S7_Optimized_Access := 'TRUE' }
VERSION : 0.1
   VAR_INPUT
      IN_tInterfaceID : Hw_Any;
      IN_tRemoteAddress : IP_V4;
      IN_tIDSend : Conn_Ouc;   // Connection ID
      IN_uiRemotePortSend : UInt;
      IN_tIDRecived : Conn_Ouc;
      IN_uiLocalPorrtRecived : UInt;
      IN_xRequestSend : Bool;
      IN_xGeneralReset : Bool;
      IN_xResetAlarm : Bool;
      IN_xThisPLCActive : Bool;
      IN_xSwitchIpInProgress : Bool;
   END_VAR
   VAR_OUTPUT
      OUT_xTSendDone : Bool;
      OUT_xTReceivedDone : Bool;
   END_VAR
   VAR_IN_OUT
      tDataToSend : Struct
         dIndexParameter : DInt;
         dByteToSend : DInt;
         rgbSendBuffer : Array[0..500] of Byte;   // FM152 - Temporary send buffer
      END_STRUCT;
      tDataRecived : Struct
         dIndexParameter : DInt;
         dByteToSend : DInt;
         rgbSendBuffer : Array[0..500] of Byte;   // FM152 - Temporary send buffer
      END_STRUCT;
   END_VAR
   VAR
      tALM : Struct   // HMI Alarms
         tS : Struct   // Stopping faults
            xErrorSendParameter : Bool;   // Error Send Parameter at BAckUp PLC
            xSpare_1 : Bool;
            xSpare_2 : Bool;
            xSpare_3 : Bool;
            xSpare_4 : Bool;
            xSpare_5 : Bool;
            xSpare_6 : Bool;
            xSpare_7 : Bool;
            xSpare_8 : Bool;
            xSpare_9 : Bool;
            xSpare_10 : Bool;
            xSpare_11 : Bool;
            xSpare_12 : Bool;
            xSpare_13 : Bool;
            xSpare_14 : Bool;
            xSpare_15 : Bool;
            xSpare_16 : Bool;
            xSpare_17 : Bool;
            xSpare_18 : Bool;
            xSpare_19 : Bool;
            xSpare_20 : Bool;
            xSpare_21 : Bool;
            xSpare_22 : Bool;
            xSpare_23 : Bool;
            xSpare_24 : Bool;
            xSpare_25 : Bool;
            xSpare_26 : Bool;
            xSpare_27 : Bool;
            xSpare_28 : Bool;
            xSpare_29 : Bool;
            xSpare_30 : Bool;
            xSpare_31 : Bool;
         END_STRUCT;
         tF : Struct   // Faults
            xSpare_0 : Bool;
            xSpare_1 : Bool;
            xSpare_2 : Bool;
            xSpare_3 : Bool;
            xSpare_4 : Bool;
            xSpare_5 : Bool;
            xSpare_6 : Bool;
            xSpare_7 : Bool;
            xSpare_8 : Bool;
            xSpare_9 : Bool;
            xSpare_10 : Bool;
            xSpare_11 : Bool;
            xSpare_12 : Bool;
            xSpare_13 : Bool;
            xSpare_14 : Bool;
            xSpare_15 : Bool;
            xSpare_16 : Bool;
            xSpare_17 : Bool;
            xSpare_18 : Bool;
            xSpare_19 : Bool;
            xSpare_20 : Bool;
            xSpare_21 : Bool;
            xSpare_22 : Bool;
            xSpare_23 : Bool;
            xSpare_24 : Bool;
            xSpare_25 : Bool;
            xSpare_26 : Bool;
            xSpare_27 : Bool;
            xSpare_28 : Bool;
            xSpare_29 : Bool;
            xSpare_30 : Bool;
            xSpare_31 : Bool;
         END_STRUCT;
         tW : Struct   // Warnings
            xSpare_0 : Bool;
            xSpare_1 : Bool;
            xSpare_2 : Bool;
            xSpare_3 : Bool;
            xSpare_4 : Bool;
            xSpare_5 : Bool;
            xSpare_6 : Bool;
            xSpare_7 : Bool;
            xSpare_8 : Bool;
            xSpare_9 : Bool;
            xSpare_10 : Bool;
            xSpare_11 : Bool;
            xSpare_12 : Bool;
            xSpare_13 : Bool;
            xSpare_14 : Bool;
            xSpare_15 : Bool;
            xSpare_16 : Bool;
            xSpare_17 : Bool;
            xSpare_18 : Bool;
            xSpare_19 : Bool;
            xSpare_20 : Bool;
            xSpare_21 : Bool;
            xSpare_22 : Bool;
            xSpare_23 : Bool;
            xSpare_24 : Bool;
            xSpare_25 : Bool;
            xSpare_26 : Bool;
            xSpare_27 : Bool;
            xSpare_28 : Bool;
            xSpare_29 : Bool;
            xSpare_30 : Bool;
            xSpare_31 : Bool;
         END_STRUCT;
      END_STRUCT;
   END_VAR
   VAR RETAIN
      tHMR : Struct
         xErrorTrasmissionParameter : Bool;   // Error trasmission parameter to PLC BackUp
         dCountSendCycle : DInt;   // Count Send Done Cycle
      END_STRUCT;
   END_VAR
   VAR
      ST_xResetSendConnection : Bool;   // FM152 - Reset the estabilished send connection
      ST_xResetRecvConnection : Bool;
      ST_xPLCActive : Bool;
      ST_xRequestActivePLC : Bool;
      ST_xRequestDeactivePLC : Bool;
      ST_xPhaseInProgress : Bool;
      OS_ReopenConnection : Bool;
      OSR_xChangeState : Bool;
      OSN_xChangeState : Bool;
      AUX_dNumByteToSend : DInt;   // FM152 - Number of byte to send
      AUX_tConnDataTSend : TCON_IP_v4;   // FM152 - Connection data structure
      AUX_tConnDataTRecive : TCON_IP_v4;   // FM152 - Connection data structure
      tPhases : Struct   // Phases
         xRequestSend : Bool;
         xEndRequestSend : Bool;
         xReqSwitchConnectPLC : Bool;
         xCloseExistinConnection : Bool;
         xReopenConnection : Bool;
         xEndSwitch : Bool;
         xSpare6 : Bool;
         xSpare7 : Bool;
         xSpare8 : Bool;
         xSpare9 : Bool;
         xSpare10 : Bool;
         xSpare11 : Bool;
         xSpare12 : Bool;
         xSpare13 : Bool;
         xSpare14 : Bool;
         xSpare15 : Bool;
         xSpare16 : Bool;
         xSpare17 : Bool;
         xSpare18 : Bool;
         xSpare19 : Bool;
         xSpare20 : Bool;
         xSpare21 : Bool;
         xSpare22 : Bool;
         xSpare23 : Bool;
         xSpare24 : Bool;
         xSpare25 : Bool;
         xSpare26 : Bool;
         xSpare27 : Bool;
         xSpare28 : Bool;
         xSpare29 : Bool;
         xSpare30 : Bool;
         xSpare31 : Bool;
      END_STRUCT;
      tmON_TimeoutSendData : TON_TIME;
      tmON_WaitConnectionClose : TON_TIME;
      tmON_WaitReopenConn : TON_TIME;
      FB_TSend : TSEND_C;
      FB_TRecv : TRCV_C;
   END_VAR
   VAR_TEMP
      TMP_dwValue : DWord;
   END_VAR
   VAR CONSTANT
      CONST_BCONNTYPE : Byte := 16#11;   // FM152 - Connection type
      CONST_DTIMEOUTSENDDATA_MS : DInt := 5000;
   END_VAR
   VAR_TEMP   // added for the SCL form of the ladder/FBD networks
      _w1 : Bool;
      _w2 : Bool;
   END_VAR
BEGIN

REGION Network 1 (SCL): Initialize connection data

           //TSend
           #AUX_tConnDataTSend.InterfaceId := #IN_tInterfaceID;
           #AUX_tConnDataTSend.ID := #IN_tIDSend;
           #AUX_tConnDataTSend.ConnectionType := #CONST_BCONNTYPE;
           #AUX_tConnDataTSend.ActiveEstablished := TRUE;
           #AUX_tConnDataTSend.RemoteAddress := #IN_tRemoteAddress;
           #AUX_tConnDataTSend.RemotePort := #IN_uiRemotePortSend;
           #AUX_tConnDataTSend.LocalPort := 0;


           //TRecived
           #AUX_tConnDataTRecive.InterfaceId := #IN_tInterfaceID;
           #AUX_tConnDataTRecive.ID := #IN_tIDRecived;
           #AUX_tConnDataTRecive.ConnectionType := #CONST_BCONNTYPE;
           #AUX_tConnDataTRecive.ActiveEstablished := False;
           #AUX_tConnDataTRecive.LocalPort := #IN_uiLocalPorrtRecived;

   IF #IN_xResetAlarm THEN
           //Reset della Allarm
           #TMP_dwValue := 0;
           SCATTER(IN := #TMP_dwValue,
                   OUT => #tALM.tS);
           #TMP_dwValue := 0;
           SCATTER(IN := #TMP_dwValue,
                   OUT => #tALM.tF);
           #TMP_dwValue := 0;
           SCATTER(IN := #TMP_dwValue,
                   OUT => #tALM.tW);
   END_IF;



   (*IF #FB_TSend.STATUS <> b#16#04 THEN
       #tPhases.xRequestSend := FALSE;
   END_IF;*)

   IF #IN_xGeneralReset THEN
           //Reset della fasi
       #TMP_dwValue := 0;
       SCATTER(IN := #TMP_dwValue,
           OUT => #tPhases);
   END_IF;


       #ST_xResetRecvConnection := #IN_xGeneralReset;
       #ST_xResetSendConnection := #IN_xGeneralReset;
END_REGION

REGION Network 2: - - - - - - - Change Connection - - - - - - --
END_REGION

REGION Network 3: Request Active or Deactive Connection
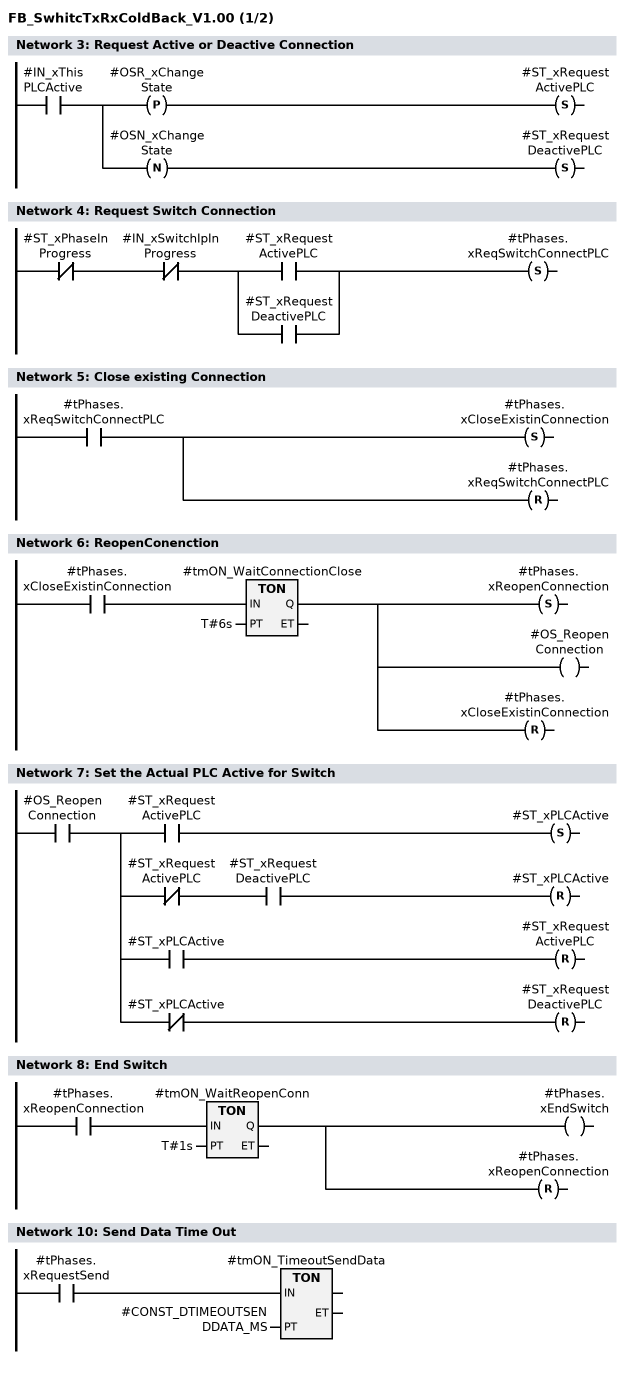
   RUNG wire#powerrail
      Contact( #IN_xThisPLCActive )
      wire#w1
      P_Trig( #OSR_xChangeState )
      S_Coil( #ST_xRequestActivePLC )
   END_RUNG
   RUNG wire#w1
      N_Trig( #OSN_xChangeState )
      S_Coil( #ST_xRequestDeactivePLC )
   END_RUNG
   // the same network as SCL:
   #_w1 := #IN_xThisPLCActive AND NOT #OSR_xChangeState;   // rising edge
   #OSR_xChangeState := #IN_xThisPLCActive;
   IF #_w1 THEN #ST_xRequestActivePLC := TRUE; END_IF;
   #_w2 := NOT #IN_xThisPLCActive AND #OSN_xChangeState;   // falling edge
   #OSN_xChangeState := #IN_xThisPLCActive;
   IF #_w2 THEN #ST_xRequestDeactivePLC := TRUE; END_IF;
END_REGION

REGION Network 4: Request Switch Connection
   RUNG wire#powerrail
      I_Contact( #ST_xPhaseInProgress )
      I_Contact( #IN_xSwitchIpInProgress )
      wire#w1
      Contact( #ST_xRequestActivePLC )
      wire#w2
      S_Coil( #tPhases.xReqSwitchConnectPLC )
   END_RUNG
   RUNG wire#w1
      Contact( #ST_xRequestDeactivePLC )
   END_RUNG wire#w2
   // the same network as SCL:
   IF NOT #ST_xPhaseInProgress AND NOT #IN_xSwitchIpInProgress AND (#ST_xRequestActivePLC OR #ST_xRequestDeactivePLC) THEN
       #tPhases.xReqSwitchConnectPLC := TRUE;
   END_IF;
END_REGION

REGION Network 5: Close existing Connection
   RUNG wire#powerrail
      Contact( #tPhases.xReqSwitchConnectPLC )
      wire#w1
      S_Coil( #tPhases.xCloseExistinConnection )
   END_RUNG
   RUNG wire#w1
      R_Coil( #tPhases.xReqSwitchConnectPLC )
   END_RUNG
   // the same network as SCL:
   IF #tPhases.xReqSwitchConnectPLC THEN
       #tPhases.xCloseExistinConnection := TRUE;
       #tPhases.xReqSwitchConnectPLC := FALSE;
   END_IF;
END_REGION

REGION Network 6: ReopenConenction
   #tmON_WaitConnectionClose(IN := #tPhases.xCloseExistinConnection, PT := T#6s);   // TON
   IF #tmON_WaitConnectionClose.Q THEN #tPhases.xReopenConnection := TRUE; END_IF;
   #OS_ReopenConnection := #tmON_WaitConnectionClose.Q;
   IF #tmON_WaitConnectionClose.Q THEN #tPhases.xCloseExistinConnection := FALSE; END_IF;
END_REGION

REGION Network 7: Set the Actual PLC Active for Switch
   RUNG wire#powerrail
      Contact( #OS_ReopenConnection )
      wire#w1
      Contact( #ST_xRequestActivePLC )
      S_Coil( #ST_xPLCActive )
   END_RUNG
   RUNG wire#w1
      I_Contact( #ST_xRequestActivePLC )
      Contact( #ST_xRequestDeactivePLC )
      R_Coil( #ST_xPLCActive )
   END_RUNG
   RUNG wire#w1
      Contact( #ST_xPLCActive )
      R_Coil( #ST_xRequestActivePLC )
   END_RUNG
   RUNG wire#w1
      I_Contact( #ST_xPLCActive )
      R_Coil( #ST_xRequestDeactivePLC )
   END_RUNG
   // the same network as SCL:
   IF #OS_ReopenConnection AND #ST_xRequestActivePLC THEN #ST_xPLCActive := TRUE; END_IF;
   IF #OS_ReopenConnection AND NOT #ST_xRequestActivePLC AND #ST_xRequestDeactivePLC THEN
       #ST_xPLCActive := FALSE;
   END_IF;
   IF #OS_ReopenConnection AND #ST_xPLCActive THEN #ST_xRequestActivePLC := FALSE; END_IF;
   IF #OS_ReopenConnection AND NOT #ST_xPLCActive THEN #ST_xRequestDeactivePLC := FALSE; END_IF;
END_REGION
